   // stn[27].wipBtn[19,7] := 129000;
   // stn[27].wipBtn[20,0] := 1000;
   // stn[27].wipBtn[20,1] := 244000;
   // stn[27].wipBtn[20,2] := 131000;
   // stn[27].wipBtn[20,3] := 1000;
   // stn[27].wipBtn[20,4] := 1000;
   // stn[27].wipBtn[20,5] := 1000;
   // stn[27].wipBtn[20,6] := 127000;
   // stn[27].wipBtn[20,7] := 132000;
   // stn[27].wipBtn[21,0] := 1000;
   // stn[27].wipBtn[21,1] := 244000;
   // stn[27].wipBtn[21,2] := 133000;
   // stn[27].wipBtn[21,3] := 1000;
   // stn[27].wipBtn[21,4] := 1000;
   // stn[27].wipBtn[21,5] := 1000;
   // stn[27].wipBtn[21,6] := 144000;
   // stn[27].wipBtn[21,7] := 134000;
   // stn[27].wipBtn[22,0] := 1000;
   // stn[27].wipBtn[22,1] := 244000;
   // stn[27].wipBtn[22,2] := 135000;
   // stn[27].wipBtn[22,3] := 1000;
   // stn[27].wipBtn[22,4] := 1000;
   // stn[27].wipBtn[22,5] := 1000;
   // stn[27].wipBtn[22,6] := 144000;
   // stn[27].wipBtn[22,7] := 136000;
   // stn[27].wipBtn[23,0] := 1000;
   // stn[27].wipBtn[23,1] := 244000;
   // stn[27].wipBtn[23,2] := 143000;
   // stn[27].wipBtn[23,3] := 1000;
   // stn[27].wipBtn[23,4] := 1000;
   // stn[27].wipBtn[23,5] := 1000;
   // stn[27].wipBtn[23,6] := 144000;
   // stn[27].wipBtn[23,7] := 134000;
   // stn[27].wipBtn[24,0] := 1000;
   // stn[27].wipBtn[24,1] := 244000;
   // stn[27].wipBtn[24,2] := 137000;
   // stn[27].wipBtn[24,3] := 1000;
   // stn[27].wipBtn[24,4] := 1000;
   // stn[27].wipBtn[24,5] := 1000;
   // stn[27].wipBtn[24,6] := 144000;
   // stn[27].wipBtn[24,7] := 136000;
   // stn[27].wipBtn[25,0] := 1000;
   // stn[27].wipBtn[25,1] := 244000;
   // stn[27].wipBtn[25,2] := 138000;
   // stn[27].wipBtn[25,3] := 1000;
   // stn[27].wipBtn[25,4] := 1000;
   // stn[27].wipBtn[25,5] := 1000;
   // stn[27].wipBtn[25,6] := 141000;
   // stn[27].wipBtn[25,7] := 129000;
   // stn[27].wipBtn[26,0] := 1000;
   // stn[27].wipBtn[26,1] := 244000;
   // stn[27].wipBtn[26,2] := 139000;
   // stn[27].wipBtn[26,3] := 1000;
   // stn[27].wipBtn[26,4] := 1000;
   // stn[27].wipBtn[26,5] := 1000;
   // stn[27].wipBtn[26,6] := 141000;
   // stn[27].wipBtn[26,7] := 140000;
   // stn[27].wipBtn[27,0] := 1000;
   // stn[27].wipBtn[27,1] := 244000;
   // stn[27].wipBtn[27,2] := 142000;
   // stn[27].wipBtn[27,3] := 1000;
   // stn[27].wipBtn[27,4] := 1000;
   // stn[27].wipBtn[27,5] := 1000;
   // stn[27].wipBtn[27,6] := 141000;
   // stn[27].wipBtn[27,7] := 126000;
   // stn[27].wipBtn[28,0] := 1000;
   // stn[27].wipBtn[28,1] := 244000;
   // stn[27].wipBtn[28,2] := 149000;
   // stn[27].wipBtn[28,3] := 1000;
   // stn[27].wipBtn[28,4] := 1000;
   // stn[27].wipBtn[28,5] := 1000;
   // stn[27].wipBtn[28,6] := 145000;
   // stn[27].wipBtn[28,7] := 150000;
   // stn[27].wipBtn[29,0] := 1000;
   // stn[27].wipBtn[29,1] := 244000;
   // stn[27].wipBtn[29,2] := 146000;
   // stn[27].wipBtn[29,3] := 1000;
   // stn[27].wipBtn[29,4] := 1000;
   // stn[27].wipBtn[29,5] := 1000;
   // stn[27].wipBtn[29,6] := 148000;
   // stn[27].wipBtn[29,7] := 147000;
   // stn[27].wipBtn[30,0] := 1000;
   // stn[27].wipBtn[30,1] := 244000;
   // stn[27].wipBtn[30,2] := 160000;
   // stn[27].wipBtn[30,3] := 1000;
   // stn[27].wipBtn[30,4] := 1000;
   // stn[27].wipBtn[30,5] := 1000;
   // stn[27].wipBtn[30,6] := 145000;
   // stn[27].wipBtn[30,7] := 161000;
   // stn[27].wipBtn[31,0] := 1000;
   // stn[27].wipBtn[31,1] := 244000;
   // stn[27].wipBtn[31,2] := 164000;
   // stn[27].wipBtn[31,3] := 1000;
   // stn[27].wipBtn[31,4] := 1000;
   // stn[27].wipBtn[31,5] := 1000;
   // stn[27].wipBtn[31,6] := 148000;
   // stn[27].wipBtn[31,7] := 147000;
   // stn[27].wipBtn[32,0] := 1000;
   // stn[27].wipBtn[32,1] := 244000;
   // stn[27].wipBtn[32,2] := 160000;
   // stn[27].wipBtn[32,3] := 1000;
   // stn[27].wipBtn[32,4] := 1000;
   // stn[27].wipBtn[32,5] := 1000;
   // stn[27].wipBtn[32,6] := 148000;
   // stn[27].wipBtn[32,7] := 161000;
   // stn[27].wipBtn[33,0] := 1000;
   // stn[27].wipBtn[33,1] := 244000;
   // stn[27].wipBtn[33,2] := 153000;
   // stn[27].wipBtn[33,3] := 152000;
   // stn[27].wipBtn[33,4] := 1000;
   // stn[27].wipBtn[33,5] := 151000;
   // stn[27].wipBtn[33,6] := 155000;
   // stn[27].wipBtn[33,7] := 154000;
   // stn[27].wipBtn[34,0] := 1000;
   // stn[27].wipBtn[34,1] := 244000;
   // stn[27].wipBtn[34,2] := 153000;
   // stn[27].wipBtn[34,3] := 1000;
   // stn[27].wipBtn[34,4] := 1000;
   // stn[27].wipBtn[34,5] := 156000;
   // stn[27].wipBtn[34,6] := 155000;
   // stn[27].wipBtn[34,7] := 154000;
   // stn[27].wipBtn[35,0] := 1000;
   // stn[27].wipBtn[35,1] := 244000;
   // stn[27].wipBtn[35,2] := 157000;
   // stn[27].wipBtn[35,3] := 1000;
   // stn[27].wipBtn[35,4] := 1000;
   // stn[27].wipBtn[35,5] := 1000;
   // stn[27].wipBtn[35,6] := 155000;
   // stn[27].wipBtn[35,7] := 158000;
   // stn[27].wipBtn[36,0] := 1000;
   // stn[27].wipBtn[36,1] := 244000;
   // stn[27].wipBtn[36,2] := 160000;
   // stn[27].wipBtn[36,3] := 1000;
   // stn[27].wipBtn[36,4] := 1000;
   // stn[27].wipBtn[36,5] := 1000;
   // stn[27].wipBtn[36,6] := 162000;
   // stn[27].wipBtn[36,7] := 161000;
   // stn[27].wipBtn[37,0] := 1000;
   // stn[27].wipBtn[37,1] := 244000;
   // stn[27].wipBtn[37,2] := 159000;
   // stn[27].wipBtn[37,3] := 1000;
   // stn[27].wipBtn[37,4] := 1000;
   // stn[27].wipBtn[37,5] := 1000;
   // stn[27].wipBtn[37,6] := 162000;
   // stn[27].wipBtn[37,7] := 161000;
   // stn[27].wipBtn[38,0] := 1000;
   // stn[27].wipBtn[38,1] := 244000;
   // stn[27].wipBtn[38,2] := 163000;
   // stn[27].wipBtn[38,3] := 1000;
   // stn[27].wipBtn[38,4] := 1000;
   // stn[27].wipBtn[38,5] := 1000;
   // stn[27].wipBtn[38,6] := 162000;
   // stn[27].wipBtn[38,7] := 161000;
   // stn[27].wipBtn[39,0] := 1000;
   // stn[27].wipBtn[39,1] := 244000;
   // stn[27].wipBtn[39,2] := 164000;
   // stn[27].wipBtn[39,3] := 1000;
   // stn[27].wipBtn[39,4] := 1000;
   // stn[27].wipBtn[39,5] := 1000;
   // stn[27].wipBtn[39,6] := 162000;
   // stn[27].wipBtn[39,7] := 147000;
   // stn[27].wipBtn[40,0] := 1000;
   // stn[27].wipBtn[40,1] := 244000;
   // stn[27].wipBtn[40,2] := 106000;
   // stn[27].wipBtn[40,3] := 129000;
   // stn[27].wipBtn[40,4] := 1000;
   // stn[27].wipBtn[40,5] := 128000;
   // stn[27].wipBtn[40,6] := 127000;
   // stn[27].wipBtn[40,7] := 134000;
   // stn[27].wipBtn[41,0] := 1000;
   // stn[27].wipBtn[41,1] := 244000;
   // stn[27].wipBtn[41,2] := 1000;
   // stn[27].wipBtn[41,3] := 1000;
   // stn[27].wipBtn[41,4] := 1000;
   // stn[27].wipBtn[41,5] := 1000;
   // stn[27].wipBtn[41,6] := 1000;
   // stn[27].wipBtn[41,7] := 1000;
   // stn[27].wipBtn[42,0] := 1000;
   // stn[27].wipBtn[42,1] := 244000;
   // stn[27].wipBtn[42,2] := 1000;
   // stn[27].wipBtn[42,3] := 1000;
   // stn[27].wipBtn[42,4] := 1000;
   // stn[27].wipBtn[42,5] := 1000;
   // stn[27].wipBtn[42,6] := 1000;
   // stn[27].wipBtn[42,7] := 1000;
   // stn[27].wipBtn[43,0] := 1000;
   // stn[27].wipBtn[43,1] := 244000;
   // stn[27].wipBtn[43,2] := 1000;
   // stn[27].wipBtn[43,3] := 1000;
   // stn[27].wipBtn[43,4] := 1000;
   // stn[27].wipBtn[43,5] := 1000;
   // stn[27].wipBtn[43,6] := 1000;
   // stn[27].wipBtn[43,7] := 1000;
   // stn[27].wipBtn[44,0] := 1000;
   // stn[27].wipBtn[44,1] := 244000;
   // stn[27].wipBtn[44,2] := 1000;
   // stn[27].wipBtn[44,3] := 1000;
   // stn[27].wipBtn[44,4] := 1000;
   // stn[27].wipBtn[44,5] := 1000;
   // stn[27].wipBtn[44,6] := 1000;
   // stn[27].wipBtn[44,7] := 1000;
   // stn[27].wipBtn[45,0] := 1000;
   // stn[27].wipBtn[45,1] := 244000;
   // stn[27].wipBtn[45,2] := 1000;
   // stn[27].wipBtn[45,3] := 1000;
   // stn[27].wipBtn[45,4] := 1000;
   // stn[27].wipBtn[45,5] := 1000;
   // stn[27].wipBtn[45,6] := 1000;
   // stn[27].wipBtn[45,7] := 1000;
   // stn[27].wipBtn[46,0] := 1000;
   // stn[27].wipBtn[46,1] := 244000;
   // stn[27].wipBtn[46,2] := 1000;
   // stn[27].wipBtn[46,3] := 1000;
   // stn[27].wipBtn[46,4] := 1000;
   // stn[27].wipBtn[46,5] := 1000;
   // stn[27].wipBtn[46,6] := 1000;
   // stn[27].wipBtn[46,7] := 1000;
   // stn[27].wipBtn[47,0] := 1000;
   // stn[27].wipBtn[47,1] := 244000;
   // stn[27].wipBtn[47,2] := 1000;
   // stn[27].wipBtn[47,3] := 1000;
   // stn[27].wipBtn[47,4] := 1000;
   // stn[27].wipBtn[47,5] := 1000;
   // stn[27].wipBtn[47,6] := 1000;
   // stn[27].wipBtn[47,7] := 1000;
   // stn[27].wipBtn[48,0] := 1000;
   // stn[27].wipBtn[48,1] := 244000;
   // stn[27].wipBtn[48,2] := 1000;
   // stn[27].wipBtn[48,3] := 1000;
   // stn[27].wipBtn[48,4] := 1000;
   // stn[27].wipBtn[48,5] := 1000;
   // stn[27].wipBtn[48,6] := 1000;
   // stn[27].wipBtn[48,7] := 1000;
   // stn[27].wipBtn[49,0] := 1000;
   // stn[27].wipBtn[49,1] := 244000;
   // stn[27].wipBtn[49,2] := 1000;
   // stn[27].wipBtn[49,3] := 1000;
   // stn[27].wipBtn[49,4] := 1000;
   // stn[27].wipBtn[49,5] := 1000;
   // stn[27].wipBtn[49,6] := 1000;
   // stn[27].wipBtn[49,7] := 1000;
   // stn[28].wipBtn[0,0] := 1000;
   // stn[28].wipBtn[0,1] := 244000;
   // stn[28].wipBtn[0,2] := 53000;
   // stn[28].wipBtn[0,3] := 1000;
   // stn[28].wipBtn[0,4] := 1000;
   // stn[28].wipBtn[0,5] := 1000;
   // stn[28].wipBtn[0,6] := 32000;
   // stn[28].wipBtn[0,7] := 74000;
   // stn[28].wipBtn[1,0] := 1000;
   // stn[28].wipBtn[1,1] := 244000;
   // stn[28].wipBtn[1,2] := 218000;
   // stn[28].wipBtn[1,3] := 1000;
   // stn[28].wipBtn[1,4] := 1000;
   // stn[28].wipBtn[1,5] := 1000;
   // stn[28].wipBtn[1,6] := 219000;
   // stn[28].wipBtn[1,7] := 224000;
   // stn[28].wipBtn[2,0] := 1000;
   // stn[28].wipBtn[2,1] := 244000;
   // stn[28].wipBtn[2,2] := 229000;
   // stn[28].wipBtn[2,3] := 232000;
   // stn[28].wipBtn[2,4] := 1000;
   // stn[28].wipBtn[2,5] := 230000;
   // stn[28].wipBtn[2,6] := 228000;
   // stn[28].wipBtn[2,7] := 231000;
   // stn[28].wipBtn[3,0] := 1000;
   // stn[28].wipBtn[3,1] := 244000;
   // stn[28].wipBtn[3,2] := 165000;
   // stn[28].wipBtn[3,3] := 1000;
   // stn[28].wipBtn[3,4] := 1000;
   // stn[28].wipBtn[3,5] := 166000;
   // stn[28].wipBtn[3,6] := 203000;
   // stn[28].wipBtn[3,7] := 204000;
   // stn[28].wipBtn[4,0] := 1000;
   // stn[28].wipBtn[4,1] := 244000;
   // stn[28].wipBtn[4,2] := 201000;
   // stn[28].wipBtn[4,3] := 1000;
   // stn[28].wipBtn[4,4] := 1000;
   // stn[28].wipBtn[4,5] := 202000;
   // stn[28].wipBtn[4,6] := 203000;
   // stn[28].wipBtn[4,7] := 204000;
   // stn[28].wipBtn[5,0] := 1000;
   // stn[28].wipBtn[5,1] := 244000;
   // stn[28].wipBtn[5,2] := 165000;
   // stn[28].wipBtn[5,3] := 1000;
   // stn[28].wipBtn[5,4] := 1000;
   // stn[28].wipBtn[5,5] := 166000;
   // stn[28].wipBtn[5,6] := 203000;
   // stn[28].wipBtn[5,7] := 204000;
   // stn[28].wipBtn[6,0] := 1000;
   // stn[28].wipBtn[6,1] := 244000;
   // stn[28].wipBtn[6,2] := 1000;
   // stn[28].wipBtn[6,3] := 186000;
   // stn[28].wipBtn[6,4] := 1000;
   // stn[28].wipBtn[6,5] := 1000;
   // stn[28].wipBtn[6,6] := 198000;
   // stn[28].wipBtn[6,7] := 180000;
   // stn[28].wipBtn[7,0] := 1000;
   // stn[28].wipBtn[7,1] := 244000;
   // stn[28].wipBtn[7,2] := 1000;
   // stn[28].wipBtn[7,3] := 200000;
   // stn[28].wipBtn[7,4] := 1000;
   // stn[28].wipBtn[7,5] := 1000;
   // stn[28].wipBtn[7,6] := 199000;
   // stn[28].wipBtn[7,7] := 179000;
   // stn[28].wipBtn[8,0] := 1000;
   // stn[28].wipBtn[8,1] := 1000;
   // stn[28].wipBtn[8,2] := 1000;
   // stn[28].wipBtn[8,3] := 1000;
   // stn[28].wipBtn[8,4] := 1000;
   // stn[28].wipBtn[8,5] := 1000;
   // stn[28].wipBtn[8,6] := 1000;
   // stn[28].wipBtn[8,7] := 1000;
   // stn[28].wipBtn[9,0] := 1000;
   // stn[28].wipBtn[9,1] := 1000;
   // stn[28].wipBtn[9,2] := 1000;
   // stn[28].wipBtn[9,3] := 1000;
   // stn[28].wipBtn[9,4] := 1000;
   // stn[28].wipBtn[9,5] := 1000;
   // stn[28].wipBtn[9,6] := 1000;
   // stn[28].wipBtn[9,7] := 1000;
   // stn[28].wipBtn[10,0] := 1000;
   // stn[28].wipBtn[10,1] := 1000;
   // stn[28].wipBtn[10,2] := 1000;
   // stn[28].wipBtn[10,3] := 1000;
   // stn[28].wipBtn[10,4] := 1000;
   // stn[28].wipBtn[10,5] := 1000;
   // stn[28].wipBtn[10,6] := 1000;
   // stn[28].wipBtn[10,7] := 1000;
   // stn[28].wipBtn[11,0] := 1000;
   // stn[28].wipBtn[11,1] := 1000;
   // stn[28].wipBtn[11,2] := 1000;
   // stn[28].wipBtn[11,3] := 1000;
   // stn[28].wipBtn[11,4] := 1000;
   // stn[28].wipBtn[11,5] := 1000;
   // stn[28].wipBtn[11,6] := 1000;
   // stn[28].wipBtn[11,7] := 1000;
   // stn[28].wipBtn[12,0] := 1000;
   // stn[28].wipBtn[12,1] := 1000;
   // stn[28].wipBtn[12,2] := 1000;
   // stn[28].wipBtn[12,3] := 1000;
   // stn[28].wipBtn[12,4] := 1000;
   // stn[28].wipBtn[12,5] := 1000;
   // stn[28].wipBtn[12,6] := 1000;
   // stn[28].wipBtn[12,7] := 1000;
   // stn[28].wipBtn[13,0] := 1000;
   // stn[28].wipBtn[13,1] := 1000;
   // stn[28].wipBtn[13,2] := 1000;
   // stn[28].wipBtn[13,3] := 1000;
   // stn[28].wipBtn[13,4] := 1000;
   // stn[28].wipBtn[13,5] := 1000;
   // stn[28].wipBtn[13,6] := 1000;
   // stn[28].wipBtn[13,7] := 1000;
   // stn[28].wipBtn[14,0] := 1000;
   // stn[28].wipBtn[14,1] := 1000;
   // stn[28].wipBtn[14,2] := 1000;
   // stn[28].wipBtn[14,3] := 1000;
   // stn[28].wipBtn[14,4] := 1000;
   // stn[28].wipBtn[14,5] := 1000;
   // stn[28].wipBtn[14,6] := 1000;
   // stn[28].wipBtn[14,7] := 1000;
   // stn[28].wipBtn[15,0] := 1000;
   // stn[28].wipBtn[15,1] := 1000;
   // stn[28].wipBtn[15,2] := 1000;
   // stn[28].wipBtn[15,3] := 1000;
   // stn[28].wipBtn[15,4] := 1000;
   // stn[28].wipBtn[15,5] := 1000;
   // stn[28].wipBtn[15,6] := 1000;
   // stn[28].wipBtn[15,7] := 1000;
   // stn[28].wipBtn[16,0] := 1000;
   // stn[28].wipBtn[16,1] := 1000;
   // stn[28].wipBtn[16,2] := 1000;
   // stn[28].wipBtn[16,3] := 1000;
   // stn[28].wipBtn[16,4] := 1000;
   // stn[28].wipBtn[16,5] := 1000;
   // stn[28].wipBtn[16,6] := 1000;
   // stn[28].wipBtn[16,7] := 1000;
   // stn[28].wipBtn[17,0] := 1000;
   // stn[28].wipBtn[17,1] := 1000;
   // stn[28].wipBtn[17,2] := 1000;
   // stn[28].wipBtn[17,3] := 1000;
   // stn[28].wipBtn[17,4] := 1000;
   // stn[28].wipBtn[17,5] := 1000;
   // stn[28].wipBtn[17,6] := 1000;
   // stn[28].wipBtn[17,7] := 1000;
   // stn[28].wipBtn[18,0] := 1000;
   // stn[28].wipBtn[18,1] := 1000;
   // stn[28].wipBtn[18,2] := 1000;
   // stn[28].wipBtn[18,3] := 1000;
   // stn[28].wipBtn[18,4] := 1000;
   // stn[28].wipBtn[18,5] := 1000;
   // stn[28].wipBtn[18,6] := 1000;
   // stn[28].wipBtn[18,7] := 1000;
   // stn[28].wipBtn[19,0] := 1000;
   // stn[28].wipBtn[19,1] := 1000;
   // stn[28].wipBtn[19,2] := 1000;
   // stn[28].wipBtn[19,3] := 1000;
   // stn[28].wipBtn[19,4] := 1000;
   // stn[28].wipBtn[19,5] := 1000;
   // stn[28].wipBtn[19,6] := 1000;
   // stn[28].wipBtn[19,7] := 1000;
   // stn[28].wipBtn[20,0] := 1000;
   // stn[28].wipBtn[20,1] := 1000;
   // stn[28].wipBtn[20,2] := 1000;
   // stn[28].wipBtn[20,3] := 1000;
   // stn[28].wipBtn[20,4] := 1000;
   // stn[28].wipBtn[20,5] := 1000;
   // stn[28].wipBtn[20,6] := 1000;
   // stn[28].wipBtn[20,7] := 1000;
   // stn[28].wipBtn[21,0] := 1000;
   // stn[28].wipBtn[21,1] := 1000;
   // stn[28].wipBtn[21,2] := 1000;
   // stn[28].wipBtn[21,3] := 1000;
   // stn[28].wipBtn[21,4] := 1000;
   // stn[28].wipBtn[21,5] := 1000;
   // stn[28].wipBtn[21,6] := 1000;
   // stn[28].wipBtn[21,7] := 1000;
   // stn[28].wipBtn[22,0] := 1000;
   // stn[28].wipBtn[22,1] := 1000;
   // stn[28].wipBtn[22,2] := 1000;
   // stn[28].wipBtn[22,3] := 1000;
   // stn[28].wipBtn[22,4] := 1000;
   // stn[28].wipBtn[22,5] := 1000;
   // stn[28].wipBtn[22,6] := 1000;
   // stn[28].wipBtn[22,7] := 1000;
   // stn[28].wipBtn[23,0] := 1000;
   // stn[28].wipBtn[23,1] := 1000;
   // stn[28].wipBtn[23,2] := 1000;
   // stn[28].wipBtn[23,3] := 1000;
   // stn[28].wipBtn[23,4] := 1000;
   // stn[28].wipBtn[23,5] := 1000;
   // stn[28].wipBtn[23,6] := 1000;
   // stn[28].wipBtn[23,7] := 1000;
   // stn[28].wipBtn[24,0] := 1000;
   // stn[28].wipBtn[24,1] := 1000;
   // stn[28].wipBtn[24,2] := 1000;
   // stn[28].wipBtn[24,3] := 1000;
   // stn[28].wipBtn[24,4] := 1000;
   // stn[28].wipBtn[24,5] := 1000;
   // stn[28].wipBtn[24,6] := 1000;
   // stn[28].wipBtn[24,7] := 1000;
   // stn[28].wipBtn[25,0] := 1000;
   // stn[28].wipBtn[25,1] := 1000;
   // stn[28].wipBtn[25,2] := 1000;
   // stn[28].wipBtn[25,3] := 1000;
   // stn[28].wipBtn[25,4] := 1000;
   // stn[28].wipBtn[25,5] := 1000;
   // stn[28].wipBtn[25,6] := 1000;
   // stn[28].wipBtn[25,7] := 1000;
   // stn[28].wipBtn[26,0] := 1000;
   // stn[28].wipBtn[26,1] := 1000;
   // stn[28].wipBtn[26,2] := 1000;
   // stn[28].wipBtn[26,3] := 1000;
   // stn[28].wipBtn[26,4] := 1000;
   // stn[28].wipBtn[26,5] := 1000;
   // stn[28].wipBtn[26,6] := 1000;
   // stn[28].wipBtn[26,7] := 1000;
   // stn[28].wipBtn[27,0] := 1000;
   // stn[28].wipBtn[27,1] := 1000;
   // stn[28].wipBtn[27,2] := 1000;
   // stn[28].wipBtn[27,3] := 1000;
   // stn[28].wipBtn[27,4] := 1000;
   // stn[28].wipBtn[27,5] := 1000;
   // stn[28].wipBtn[27,6] := 1000;
   // stn[28].wipBtn[27,7] := 1000;
   // stn[28].wipBtn[28,0] := 1000;
   // stn[28].wipBtn[28,1] := 1000;
   // stn[28].wipBtn[28,2] := 1000;
   // stn[28].wipBtn[28,3] := 1000;
   // stn[28].wipBtn[28,4] := 1000;
   // stn[28].wipBtn[28,5] := 1000;
   // stn[28].wipBtn[28,6] := 1000;
   // stn[28].wipBtn[28,7] := 1000;
   // stn[28].wipBtn[29,0] := 1000;
   // stn[28].wipBtn[29,1] := 1000;
   // stn[28].wipBtn[29,2] := 1000;
   // stn[28].wipBtn[29,3] := 1000;
   // stn[28].wipBtn[29,4] := 1000;
   // stn[28].wipBtn[29,5] := 1000;
   // stn[28].wipBtn[29,6] := 1000;
   // stn[28].wipBtn[29,7] := 1000;
   // stn[28].wipBtn[30,0] := 1000;
   // stn[28].wipBtn[30,1] := 1000;
   // stn[28].wipBtn[30,2] := 1000;
   // stn[28].wipBtn[30,3] := 1000;
   // stn[28].wipBtn[30,4] := 1000;
   // stn[28].wipBtn[30,5] := 1000;
   // stn[28].wipBtn[30,6] := 1000;
   // stn[28].wipBtn[30,7] := 1000;
   // stn[28].wipBtn[31,0] := 1000;
   // stn[28].wipBtn[31,1] := 1000;
   // stn[28].wipBtn[31,2] := 1000;
   // stn[28].wipBtn[31,3] := 1000;
   // stn[28].wipBtn[31,4] := 1000;
   // stn[28].wipBtn[31,5] := 1000;
   // stn[28].wipBtn[31,6] := 1000;
   // stn[28].wipBtn[31,7] := 1000;
   // stn[28].wipBtn[32,0] := 1000;
   // stn[28].wipBtn[32,1] := 1000;
   // stn[28].wipBtn[32,2] := 1000;
   // stn[28].wipBtn[32,3] := 1000;
   // stn[28].wipBtn[32,4] := 1000;
   // stn[28].wipBtn[32,5] := 1000;
   // stn[28].wipBtn[32,6] := 1000;
   // stn[28].wipBtn[32,7] := 1000;
   // stn[28].wipBtn[33,0] := 1000;
   // stn[28].wipBtn[33,1] := 1000;
   // stn[28].wipBtn[33,2] := 1000;
   // stn[28].wipBtn[33,3] := 1000;
   // stn[28].wipBtn[33,4] := 1000;
   // stn[28].wipBtn[33,5] := 1000;
   // stn[28].wipBtn[33,6] := 1000;
   // stn[28].wipBtn[33,7] := 1000;
   // stn[28].wipBtn[34,0] := 1000;
   // stn[28].wipBtn[34,1] := 1000;
   // stn[28].wipBtn[34,2] := 1000;
   // stn[28].wipBtn[34,3] := 1000;
   // stn[28].wipBtn[34,4] := 1000;
   // stn[28].wipBtn[34,5] := 1000;
   // stn[28].wipBtn[34,6] := 1000;
   // stn[28].wipBtn[34,7] := 1000;
   // stn[28].wipBtn[35,0] := 1000;
   // stn[28].wipBtn[35,1] := 1000;
   // stn[28].wipBtn[35,2] := 1000;
   // stn[28].wipBtn[35,3] := 1000;
   // stn[28].wipBtn[35,4] := 1000;
   // stn[28].wipBtn[35,5] := 1000;
   // stn[28].wipBtn[35,6] := 1000;
   // stn[28].wipBtn[35,7] := 1000;
   // stn[28].wipBtn[36,0] := 1000;
   // stn[28].wipBtn[36,1] := 1000;
   // stn[28].wipBtn[36,2] := 1000;
   // stn[28].wipBtn[36,3] := 1000;
   // stn[28].wipBtn[36,4] := 1000;
   // stn[28].wipBtn[36,5] := 1000;
   // stn[28].wipBtn[36,6] := 1000;
   // stn[28].wipBtn[36,7] := 1000;
   // stn[28].wipBtn[37,0] := 1000;
   // stn[28].wipBtn[37,1] := 1000;
   // stn[28].wipBtn[37,2] := 1000;
   // stn[28].wipBtn[37,3] := 1000;
   // stn[28].wipBtn[37,4] := 1000;
   // stn[28].wipBtn[37,5] := 1000;
   // stn[28].wipBtn[37,6] := 1000;
   // stn[28].wipBtn[37,7] := 1000;
   // stn[28].wipBtn[38,0] := 1000;
   // stn[28].wipBtn[38,1] := 1000;
   // stn[28].wipBtn[38,2] := 1000;
   // stn[28].wipBtn[38,3] := 1000;
   // stn[28].wipBtn[38,4] := 1000;
   // stn[28].wipBtn[38,5] := 1000;
   // stn[28].wipBtn[38,6] := 1000;
   // stn[28].wipBtn[38,7] := 1000;
   // stn[28].wipBtn[39,0] := 1000;
   // stn[28].wipBtn[39,1] := 1000;
   // stn[28].wipBtn[39,2] := 1000;
   // stn[28].wipBtn[39,3] := 1000;
   // stn[28].wipBtn[39,4] := 1000;
   // stn[28].wipBtn[39,5] := 1000;
   // stn[28].wipBtn[39,6] := 1000;
   // stn[28].wipBtn[39,7] := 1000;
   // stn[28].wipBtn[40,0] := 1000;
   // stn[28].wipBtn[40,1] := 1000;
   // stn[28].wipBtn[40,2] := 1000;
   // stn[28].wipBtn[40,3] := 1000;
   // stn[28].wipBtn[40,4] := 1000;
   // stn[28].wipBtn[40,5] := 1000;
   // stn[28].wipBtn[40,6] := 1000;
   // stn[28].wipBtn[40,7] := 1000;
   // stn[28].wipBtn[41,0] := 1000;
   // stn[28].wipBtn[41,1] := 1000;
   // stn[28].wipBtn[41,2] := 1000;
   // stn[28].wipBtn[41,3] := 1000;
   // stn[28].wipBtn[41,4] := 1000;
   // stn[28].wipBtn[41,5] := 1000;
   // stn[28].wipBtn[41,6] := 1000;
   // stn[28].wipBtn[41,7] := 1000;
   // stn[28].wipBtn[42,0] := 1000;
   // stn[28].wipBtn[42,1] := 1000;
   // stn[28].wipBtn[42,2] := 1000;
   // stn[28].wipBtn[42,3] := 1000;
   // stn[28].wipBtn[42,4] := 1000;
   // stn[28].wipBtn[42,5] := 1000;
   // stn[28].wipBtn[42,6] := 1000;
   // stn[28].wipBtn[42,7] := 1000;
   // stn[28].wipBtn[43,0] := 1000;
   // stn[28].wipBtn[43,1] := 1000;
   // stn[28].wipBtn[43,2] := 1000;
   // stn[28].wipBtn[43,3] := 1000;
   // stn[28].wipBtn[43,4] := 1000;
   // stn[28].wipBtn[43,5] := 1000;
   // stn[28].wipBtn[43,6] := 1000;
   // stn[28].wipBtn[43,7] := 1000;
   // stn[28].wipBtn[44,0] := 1000;
   // stn[28].wipBtn[44,1] := 1000;
   // stn[28].wipBtn[44,2] := 1000;
   // stn[28].wipBtn[44,3] := 1000;
   // stn[28].wipBtn[44,4] := 1000;
   // stn[28].wipBtn[44,5] := 1000;
   // stn[28].wipBtn[44,6] := 1000;
   // stn[28].wipBtn[44,7] := 1000;
   // stn[28].wipBtn[45,0] := 1000;
   // stn[28].wipBtn[45,1] := 1000;
   // stn[28].wipBtn[45,2] := 1000;
   // stn[28].wipBtn[45,3] := 1000;
   // stn[28].wipBtn[45,4] := 1000;
   // stn[28].wipBtn[45,5] := 1000;
   // stn[28].wipBtn[45,6] := 1000;
   // stn[28].wipBtn[45,7] := 1000;
   // stn[28].wipBtn[46,0] := 1000;
   // stn[28].wipBtn[46,1] := 1000;
   // stn[28].wipBtn[46,2] := 1000;
   // stn[28].wipBtn[46,3] := 1000;
   // stn[28].wipBtn[46,4] := 1000;
   // stn[28].wipBtn[46,5] := 1000;
   // stn[28].wipBtn[46,6] := 1000;
   // stn[28].wipBtn[46,7] := 1000;
   // stn[28].wipBtn[47,0] := 1000;
   // stn[28].wipBtn[47,1] := 1000;
   // stn[28].wipBtn[47,2] := 1000;
   // stn[28].wipBtn[47,3] := 1000;
   // stn[28].wipBtn[47,4] := 1000;
   // stn[28].wipBtn[47,5] := 1000;
   // stn[28].wipBtn[47,6] := 1000;
   // stn[28].wipBtn[47,7] := 1000;
   // stn[28].wipBtn[48,0] := 1000;
   // stn[28].wipBtn[48,1] := 1000;
   // stn[28].wipBtn[48,2] := 1000;
   // stn[28].wipBtn[48,3] := 1000;
   // stn[28].wipBtn[48,4] := 1000;
   // stn[28].wipBtn[48,5] := 1000;
   // stn[28].wipBtn[48,6] := 1000;
   // stn[28].wipBtn[48,7] := 1000;
   // stn[28].wipBtn[49,0] := 1000;
   // stn[28].wipBtn[49,1] := 1000;
   // stn[28].wipBtn[49,2] := 1000;
   // stn[28].wipBtn[49,3] := 1000;
   // stn[28].wipBtn[49,4] := 1000;
   // stn[28].wipBtn[49,5] := 1000;
   // stn[28].wipBtn[49,6] := 1000;
   // stn[28].wipBtn[49,7] := 1000;
   // stn[29].wipBtn[0,0] := 1000;
   // stn[29].wipBtn[0,1] := 244000;
   // stn[29].wipBtn[0,2] := 1000;
   // stn[29].wipBtn[0,3] := 4000;
   // stn[29].wipBtn[0,4] := 1000;
   // stn[29].wipBtn[0,5] := 1000;
   // stn[29].wipBtn[0,6] := 2000;
   // stn[29].wipBtn[0,7] := 3000;
   // stn[29].wipBtn[1,0] := 1000;
   // stn[29].wipBtn[1,1] := 244000;
   // stn[29].wipBtn[1,2] := 6000;
   // stn[29].wipBtn[1,3] := 10000;
   // stn[29].wipBtn[1,4] := 1000;
   // stn[29].wipBtn[1,5] := 7000;
   // stn[29].wipBtn[1,6] := 5000;
   // stn[29].wipBtn[1,7] := 11000;
   // stn[29].wipBtn[2,0] := 1000;
   // stn[29].wipBtn[2,1] := 244000;
   // stn[29].wipBtn[2,2] := 8000;
   // stn[29].wipBtn[2,3] := 10000;
   // stn[29].wipBtn[2,4] := 1000;
   // stn[29].wipBtn[2,5] := 9000;
   // stn[29].wipBtn[2,6] := 5000;
   // stn[29].wipBtn[2,7] := 11000;
   // stn[29].wipBtn[3,0] := 1000;
   // stn[29].wipBtn[3,1] := 1000;
   // stn[29].wipBtn[3,2] := 1000;
   // stn[29].wipBtn[3,3] := 1000;
   // stn[29].wipBtn[3,4] := 1000;
   // stn[29].wipBtn[3,5] := 1000;
   // stn[29].wipBtn[3,6] := 1000;
   // stn[29].wipBtn[3,7] := 1000;
   // stn[29].wipBtn[4,0] := 1000;
   // stn[29].wipBtn[4,1] := 1000;
   // stn[29].wipBtn[4,2] := 1000;
   // stn[29].wipBtn[4,3] := 1000;
   // stn[29].wipBtn[4,4] := 1000;
   // stn[29].wipBtn[4,5] := 1000;
   // stn[29].wipBtn[4,6] := 1000;
   // stn[29].wipBtn[4,7] := 1000;
   // stn[29].wipBtn[5,0] := 1000;
   // stn[29].wipBtn[5,1] := 1000;
   // stn[29].wipBtn[5,2] := 1000;
   // stn[29].wipBtn[5,3] := 1000;
   // stn[29].wipBtn[5,4] := 1000;
   // stn[29].wipBtn[5,5] := 1000;
   // stn[29].wipBtn[5,6] := 1000;
   // stn[29].wipBtn[5,7] := 1000;
   // stn[29].wipBtn[6,0] := 1000;
   // stn[29].wipBtn[6,1] := 1000;
   // stn[29].wipBtn[6,2] := 1000;
   // stn[29].wipBtn[6,3] := 1000;
   // stn[29].wipBtn[6,4] := 1000;
   // stn[29].wipBtn[6,5] := 1000;
   // stn[29].wipBtn[6,6] := 1000;
   // stn[29].wipBtn[6,7] := 1000;
   // stn[29].wipBtn[7,0] := 1000;
   // stn[29].wipBtn[7,1] := 1000;
   // stn[29].wipBtn[7,2] := 1000;
   // stn[29].wipBtn[7,3] := 1000;
   // stn[29].wipBtn[7,4] := 1000;
   // stn[29].wipBtn[7,5] := 1000;
   // stn[29].wipBtn[7,6] := 1000;
   // stn[29].wipBtn[7,7] := 1000;
   // stn[29].wipBtn[8,0] := 1000;
   // stn[29].wipBtn[8,1] := 1000;
   // stn[29].wipBtn[8,2] := 1000;
   // stn[29].wipBtn[8,3] := 1000;
   // stn[29].wipBtn[8,4] := 1000;
   // stn[29].wipBtn[8,5] := 1000;
   // stn[29].wipBtn[8,6] := 1000;
   // stn[29].wipBtn[8,7] := 1000;
   // stn[29].wipBtn[9,0] := 1000;
   // stn[29].wipBtn[9,1] := 1000;
   // stn[29].wipBtn[9,2] := 1000;
   // stn[29].wipBtn[9,3] := 1000;
   // stn[29].wipBtn[9,4] := 1000;
   // stn[29].wipBtn[9,5] := 1000;
   // stn[29].wipBtn[9,6] := 1000;
   // stn[29].wipBtn[9,7] := 1000;
   // stn[29].wipBtn[10,0] := 1000;
   // stn[29].wipBtn[10,1] := 1000;
   // stn[29].wipBtn[10,2] := 1000;
   // stn[29].wipBtn[10,3] := 1000;
   // stn[29].wipBtn[10,4] := 1000;
   // stn[29].wipBtn[10,5] := 1000;
   // stn[29].wipBtn[10,6] := 1000;
   // stn[29].wipBtn[10,7] := 1000;
   // stn[29].wipBtn[11,0] := 1000;
   // stn[29].wipBtn[11,1] := 1000;
   // stn[29].wipBtn[11,2] := 1000;
   // stn[29].wipBtn[11,3] := 1000;
   // stn[29].wipBtn[11,4] := 1000;
   // stn[29].wipBtn[11,5] := 1000;
   // stn[29].wipBtn[11,6] := 1000;
   // stn[29].wipBtn[11,7] := 1000;
   // stn[29].wipBtn[12,0] := 1000;
   // stn[29].wipBtn[12,1] := 1000;
   // stn[29].wipBtn[12,2] := 1000;
   // stn[29].wipBtn[12,3] := 1000;
   // stn[29].wipBtn[12,4] := 1000;
   // stn[29].wipBtn[12,5] := 1000;
   // stn[29].wipBtn[12,6] := 1000;
   // stn[29].wipBtn[12,7] := 1000;
   // stn[29].wipBtn[13,0] := 1000;
   // stn[29].wipBtn[13,1] := 1000;
   // stn[29].wipBtn[13,2] := 1000;
   // stn[29].wipBtn[13,3] := 1000;
   // stn[29].wipBtn[13,4] := 1000;
   // stn[29].wipBtn[13,5] := 1000;
   // stn[29].wipBtn[13,6] := 1000;
   // stn[29].wipBtn[13,7] := 1000;
   // stn[29].wipBtn[14,0] := 1000;
   // stn[29].wipBtn[14,1] := 1000;
   // stn[29].wipBtn[14,2] := 1000;
   // stn[29].wipBtn[14,3] := 1000;
   // stn[29].wipBtn[14,4] := 1000;
   // stn[29].wipBtn[14,5] := 1000;
   // stn[29].wipBtn[14,6] := 1000;
   // stn[29].wipBtn[14,7] := 1000;
   // stn[29].wipBtn[15,0] := 1000;
   // stn[29].wipBtn[15,1] := 1000;
   // stn[29].wipBtn[15,2] := 1000;
   // stn[29].wipBtn[15,3] := 1000;
   // stn[29].wipBtn[15,4] := 1000;
   // stn[29].wipBtn[15,5] := 1000;
   // stn[29].wipBtn[15,6] := 1000;
   // stn[29].wipBtn[15,7] := 1000;
   // stn[29].wipBtn[16,0] := 1000;
   // stn[29].wipBtn[16,1] := 1000;
   // stn[29].wipBtn[16,2] := 1000;
   // stn[29].wipBtn[16,3] := 1000;
   // stn[29].wipBtn[16,4] := 1000;
   // stn[29].wipBtn[16,5] := 1000;
   // stn[29].wipBtn[16,6] := 1000;
   // stn[29].wipBtn[16,7] := 1000;
   // stn[29].wipBtn[17,0] := 1000;
   // stn[29].wipBtn[17,1] := 1000;
   // stn[29].wipBtn[17,2] := 1000;
   // stn[29].wipBtn[17,3] := 1000;
   // stn[29].wipBtn[17,4] := 1000;
   // stn[29].wipBtn[17,5] := 1000;
   // stn[29].wipBtn[17,6] := 1000;
   // stn[29].wipBtn[17,7] := 1000;
   // stn[29].wipBtn[18,0] := 1000;
   // stn[29].wipBtn[18,1] := 1000;
   // stn[29].wipBtn[18,2] := 1000;
   // stn[29].wipBtn[18,3] := 1000;
   // stn[29].wipBtn[18,4] := 1000;
   // stn[29].wipBtn[18,5] := 1000;
   // stn[29].wipBtn[18,6] := 1000;
   // stn[29].wipBtn[18,7] := 1000;
   // stn[29].wipBtn[19,0] := 1000;
   // stn[29].wipBtn[19,1] := 1000;
   // stn[29].wipBtn[19,2] := 1000;
   // stn[29].wipBtn[19,3] := 1000;
   // stn[29].wipBtn[19,4] := 1000;
   // stn[29].wipBtn[19,5] := 1000;
   // stn[29].wipBtn[19,6] := 1000;
   // stn[29].wipBtn[19,7] := 1000;
   // stn[29].wipBtn[20,0] := 1000;
   // stn[29].wipBtn[20,1] := 1000;
   // stn[29].wipBtn[20,2] := 1000;
   // stn[29].wipBtn[20,3] := 1000;
   // stn[29].wipBtn[20,4] := 1000;
   // stn[29].wipBtn[20,5] := 1000;
   // stn[29].wipBtn[20,6] := 1000;
   // stn[29].wipBtn[20,7] := 1000;
   // stn[29].wipBtn[21,0] := 1000;
   // stn[29].wipBtn[21,1] := 1000;
   // stn[29].wipBtn[21,2] := 1000;
   // stn[29].wipBtn[21,3] := 1000;
   // stn[29].wipBtn[21,4] := 1000;
   // stn[29].wipBtn[21,5] := 1000;
   // stn[29].wipBtn[21,6] := 1000;
   // stn[29].wipBtn[21,7] := 1000;
   // stn[29].wipBtn[22,0] := 1000;
   // stn[29].wipBtn[22,1] := 1000;
   // stn[29].wipBtn[22,2] := 1000;
   // stn[29].wipBtn[22,3] := 1000;
   // stn[29].wipBtn[22,4] := 1000;
   // stn[29].wipBtn[22,5] := 1000;
   // stn[29].wipBtn[22,6] := 1000;
   // stn[29].wipBtn[22,7] := 1000;
   // stn[29].wipBtn[23,0] := 1000;
   // stn[29].wipBtn[23,1] := 1000;
   // stn[29].wipBtn[23,2] := 1000;
   // stn[29].wipBtn[23,3] := 1000;
   // stn[29].wipBtn[23,4] := 1000;
   // stn[29].wipBtn[23,5] := 1000;
   // stn[29].wipBtn[23,6] := 1000;
   // stn[29].wipBtn[23,7] := 1000;
   // stn[29].wipBtn[24,0] := 1000;
   // stn[29].wipBtn[24,1] := 1000;
   // stn[29].wipBtn[24,2] := 1000;
   // stn[29].wipBtn[24,3] := 1000;
   // stn[29].wipBtn[24,4] := 1000;
   // stn[29].wipBtn[24,5] := 1000;
   // stn[29].wipBtn[24,6] := 1000;
   // stn[29].wipBtn[24,7] := 1000;
   // stn[29].wipBtn[25,0] := 1000;
   // stn[29].wipBtn[25,1] := 1000;
   // stn[29].wipBtn[25,2] := 1000;
   // stn[29].wipBtn[25,3] := 1000;
   // stn[29].wipBtn[25,4] := 1000;
   // stn[29].wipBtn[25,5] := 1000;
   // stn[29].wipBtn[25,6] := 1000;
   // stn[29].wipBtn[25,7] := 1000;
   // stn[29].wipBtn[26,0] := 1000;
   // stn[29].wipBtn[26,1] := 1000;
   // stn[29].wipBtn[26,2] := 1000;
   // stn[29].wipBtn[26,3] := 1000;
   // stn[29].wipBtn[26,4] := 1000;
   // stn[29].wipBtn[26,5] := 1000;
   // stn[29].wipBtn[26,6] := 1000;
   // stn[29].wipBtn[26,7] := 1000;
   // stn[29].wipBtn[27,0] := 1000;
   // stn[29].wipBtn[27,1] := 1000;
   // stn[29].wipBtn[27,2] := 1000;
   // stn[29].wipBtn[27,3] := 1000;
   // stn[29].wipBtn[27,4] := 1000;
   // stn[29].wipBtn[27,5] := 1000;
   // stn[29].wipBtn[27,6] := 1000;
   // stn[29].wipBtn[27,7] := 1000;
   // stn[29].wipBtn[28,0] := 1000;
   // stn[29].wipBtn[28,1] := 1000;
   // stn[29].wipBtn[28,2] := 1000;
   // stn[29].wipBtn[28,3] := 1000;
   // stn[29].wipBtn[28,4] := 1000;
   // stn[29].wipBtn[28,5] := 1000;
   // stn[29].wipBtn[28,6] := 1000;
   // stn[29].wipBtn[28,7] := 1000;
   // stn[29].wipBtn[29,0] := 1000;
   // stn[29].wipBtn[29,1] := 1000;
   // stn[29].wipBtn[29,2] := 1000;
   // stn[29].wipBtn[29,3] := 1000;
   // stn[29].wipBtn[29,4] := 1000;
   // stn[29].wipBtn[29,5] := 1000;
   // stn[29].wipBtn[29,6] := 1000;
   // stn[29].wipBtn[29,7] := 1000;
   // stn[29].wipBtn[30,0] := 1000;
   // stn[29].wipBtn[30,1] := 1000;
   // stn[29].wipBtn[30,2] := 1000;
   // stn[29].wipBtn[30,3] := 1000;
   // stn[29].wipBtn[30,4] := 1000;
   // stn[29].wipBtn[30,5] := 1000;
   // stn[29].wipBtn[30,6] := 1000;
   // stn[29].wipBtn[30,7] := 1000;
   // stn[29].wipBtn[31,0] := 1000;
   // stn[29].wipBtn[31,1] := 1000;
   // stn[29].wipBtn[31,2] := 1000;
   // stn[29].wipBtn[31,3] := 1000;
   // stn[29].wipBtn[31,4] := 1000;
   // stn[29].wipBtn[31,5] := 1000;
   // stn[29].wipBtn[31,6] := 1000;
   // stn[29].wipBtn[31,7] := 1000;
   // stn[29].wipBtn[32,0] := 1000;
   // stn[29].wipBtn[32,1] := 1000;
   // stn[29].wipBtn[32,2] := 1000;
   // stn[29].wipBtn[32,3] := 1000;
   // stn[29].wipBtn[32,4] := 1000;
   // stn[29].wipBtn[32,5] := 1000;
   // stn[29].wipBtn[32,6] := 1000;
   // stn[29].wipBtn[32,7] := 1000;
   // stn[29].wipBtn[33,0] := 1000;
   // stn[29].wipBtn[33,1] := 1000;
   // stn[29].wipBtn[33,2] := 1000;
   // stn[29].wipBtn[33,3] := 1000;
   // stn[29].wipBtn[33,4] := 1000;
   // stn[29].wipBtn[33,5] := 1000;
   // stn[29].wipBtn[33,6] := 1000;
   // stn[29].wipBtn[33,7] := 1000;
   // stn[29].wipBtn[34,0] := 1000;
   // stn[29].wipBtn[34,1] := 1000;
   // stn[29].wipBtn[34,2] := 1000;
   // stn[29].wipBtn[34,3] := 1000;
   // stn[29].wipBtn[34,4] := 1000;
   // stn[29].wipBtn[34,5] := 1000;
   // stn[29].wipBtn[34,6] := 1000;
   // stn[29].wipBtn[34,7] := 1000;